// Mitsubishi GX Works2 project: KotelnyaPLC   PLC: FX3U/FX3UC
// Kotelnya

// global labels: Global1
VAR_GLOBAL
  Pw_in_K1 AT D116 : REAL;  (* Давление воды на входе в котел № 1 *)
  TwP_K1 AT D100 : REAL;  (* Температура прямой воды котел № 1 *)
  TwO_K1 AT D102 : REAL;  (* Температура обратной воды котел № 1 *)
  TwP_K2 AT D104 : REAL;  (* Температура прямой воды котел № 2 *)
  TwO_K2 AT D106 : REAL;  (* Температура обратной воды котел № 2 *)
  pusk : BOOL;  (* Переключение вывода данных в градусах "С или "F из блока Fx3U-4AD-PT-ADP *)
  Pw_out_K1 AT D114 : REAL;  (* Давление воды на выходе из котла № 1 *)
  Pw_in_K2 AT D120 : REAL;  (* Давление воды на входе в котел № 2 *)
  Pw_out_K2 AT D118 : REAL;  (* Давление воды на выходе из котла № 2 *)
  TwP AT D108 : REAL;  (* Температура сетевой воды прямой *)
  TwO AT D110 : REAL;  (* Температура сетевой воды обратной *)
  TN_air AT D112 : REAL;  (* Температура наружнего воздуха *)
  F_GAZ AT M144 : BOOL;  (* Флаг активации газового клапана *)
  F_CO_LEVEL2 AT M102 : BOOL;  (* Флаг Активация концентрации по окиси углерода выше 100МГ/М3 Порог 2 *)
  F_CO_LEVEL1 AT M101 : BOOL;  (* Флаг Активация концентрации по окиси углерода выше 20МГ/М3 Порог 1 *)
  F_CH4_LEVEL1 AT M103 : BOOL;  (* Вход Загазованность по метану 0.5% Порог 1 *)
  F_CH4_LEVEL2 AT M104 : BOOL;  (* Вход Загазованность по метану 1% Порог 2 *)
  F_FIRE_RELAY AT M105 : BOOL;  (* Флаг Входа реле пожара *)
  F_HIGH_PRESSURE_GAS AT M146 : BOOL;  (* Флаг Повышение давления газа на вводе *)
  F_LOW_PRESSURE_GAS AT M145 : BOOL;  (* Флаг Понижение давления газа на вводе *)
  F_SB6_SIGNAL_TEST : BOOL;  (* Флаг Тестирование звкового сигнала *)
  F_SB5_SOUND_OFF : BOOL;  (* Флаг Отключение звкового сигнала *)
  F_SA4_SOUND_ON : BOOL;  (* Вход- Переключатель в положении - Звуковой сигнал порога 2 включен *)
  F_SOUND_OFF : BOOL;  (* Флаг Отключение звукового сигнала *)
  F_SOUND : BOOL;  (* Флаг Активация выхода звуковой сигнал *)
  F_LOW_PRESSURE_BACKWATER AT M106 : BOOL;  (* Флаг Понижение давления обратной сетевой воды (унитерм) *)
  F_ALARM_GOR_KOTEL_1 AT M107 : BOOL;  (* Флаг авария Котла 1 *)
  F_ALARM_GOR_KOTEL_2 AT M108 : BOOL;  (* Флаг авария Котла 2 *)
  F_REZERV_PUMP_ON AT M142 : BOOL;  (* Флаг Включился резервный циркуляционный насос. Провод 325 *)
  F_SB1_KOTEL_ON : BOOL;  (* Флаг Кнопка Включения работы Котлов *)
  F_SB2_KOTEL_OFF : BOOL;  (* Флаг Кнопка Выключения работы Котлов *)
  F_SA3_KOTEL_1 : BOOL;  (* Флаг Переключение Котел 1 основной 2 резервный *)
  F_SA3_KOTEL_2 : BOOL;  (* Флаг Переключение Котел 2 основной 1 резервный *)
  F_ROTATION_B_VALVE_COOL AT M201 : BOOL;  (* Флаг Вращение трехходового клапана по часовой стрелке *)
  F_ROTATION_F_VALVE_HEAT AT M202 : BOOL;  (* Флаг Вращение трехходового клапана против часовой стрелки *)
  F_TERMOMETR_95C_KOTEL_1 AT M111 : BOOL;  (* Флаг Термометр манометрический Котел 1. 95С постоянный *)
  F_TERMOMETR_95C_KOTEL_2 AT M112 : BOOL;  (* Флаг Термометр манометрический Котел 2. 95С постоянный *)
  F_SA2_RECIRC_PUMP_1 : BOOL;  (* Флаг. Переключение Рециркуляционный насос 1, Положение Дист *)
  F_SA1_RECIRC_PUMP_1 : BOOL;  (* Флаг. Переключение Рециркуляционный насос 2, Положение Дист *)
  PwP AT D122 : REAL;  (* Давление прямой сетевой воды *)
  PwO AT D124 : REAL;  (* Давление обратной сетевой воды *)
  OP_PwO_ust AT D202 : REAL;  (* ОП Уставка обратного сетевого давления *)
  FB_KOTEL_1 : KOTEL;
  F_KOTEL_1_DOP AT M132 : BOOL;  (* Флаг Котел 1 работает в качестве дополнительного *)
  F_KOTEL_2_DOP AT M134 : BOOL;  (* Флаг Котел 2 работает в качестве дополнительного *)
  F_ALARM_KOTEL_1 AT M135 : BOOL;  (* Флаг Авария Котел 1 *)
  F_ALARM_KOTEL_2 AT M136 : BOOL;  (* Флаг Авария Котел 2 *)
  F_TERMOMETR_90C_KOTEL_1 AT M109 : BOOL;  (* Флаг Термометр манометрический Котел 1. 86С регулируемый *)
  F_TERMOMETR_90C_KOTEL_2 AT M110 : BOOL;  (* Флаг Термометр манометрический Котел 2. 86С регулируемый *)
  OP_PwMAX_ust AT D204 : REAL;  (* Давление воды максимальное Котел *)
  OP_PwMIN_ust AT D206 : REAL;  (* Давление воды минимальное Котел *)
  F_Pdn40_KOTEL_1 AT M113 : BOOL;  (* Флаг Датчик давления в топке ДН-40 Котел 1 *)
  F_Pdn40_KOTEL_2 AT M114 : BOOL;  (* Флаг Датчик давления в топке ДН-40 Котел 2 *)
  OP_Tw80_ust AT D208 : REAL;  (* Панель оператора температура большого горения *)
  OP_Tw86_ust AT D210 : REAL;  (* Панель оператора температура малого горения *)
  F_BURNER_1_KOTEL_1 AT M123 : BOOL;  (* Флаг Горелка 1 Котел 1 *)
  F_BURNER_2_KOTEL_1 AT M124 : BOOL;  (* Флаг Горелка 2 Котел 1 *)
  F_BURNER_1_KOTEL_2 AT M125 : BOOL;  (* Флаг Горелка 1 Котел 2 *)
  F_BURNER_2_KOTEL_2 AT M126 : BOOL;  (* Флаг Горелка 2 Котел 2 *)
  F_CIRC_PUMP_1 AT M140 : BOOL;  (* Флаг Включен циркуляционный насос 1 *)
  F_CIRC_PUMP_2 AT M141 : BOOL;  (* Флаг Включен циркуляционный насос 2 *)
  F_CIRC_PUMP_ON AT M116 : BOOL;  (* Включен циркуляционный насос *)
  F_RECIRC_PUMP_1 AT M127 : BOOL;  (* Флаг активации насоса рециркуляции 1 *)
  F_RECIRC_PUMP_2 AT M128 : BOOL;  (* Флаг активации насоса рециркуляции 2 *)
  OP_RST_ALARM AT M115 : BOOL;  (* Панель оператора Сброс аварии *)
  OP_Tw90_ust AT D212 : REAL;  (* Панель оператора Температура на выходе котла при которой авария *)
  TWO_ust AT D126 : REAL;  (* Температура сетевой воды обратной табличная *)
  OP_GRAPH_N AT D216 : INT;  (* Панель оператора Номер графика нагрева *)
  OP_DAY AT D200 : INT;  (* Панель оператора День *)
  OP_NIGHT AT D201 : INT;  (* Панель оператора Ночь *)
  OP_Tw65_ust AT D214 : REAL;  (* Панель оператора Температура включения рециркуляционного насоса *)
  GRAPH_1 : GRAPH;  (* FBD график определения заданной воды *)
  F_HOUR AT D128 : INT;  (* Час текущий *)
  F_MINUTE AT D129 : INT;  (* Минуты текущие *)
  F_MOTOR_RECIRC_PUMP_1 AT M121 : BOOL;  (* Флаг включен мотор-автомат рециркуляционного насоса 1 *)
  F_MOTOR_RECIRC_PUMP_2 AT M122 : BOOL;  (* Флаг включен мотор-автомат рециркуляционного насоса 2 *)
  F_KOTEL_2 AT M133 : BOOL;  (* Флаг Котел 2 *)
  F_KOTEL_1 AT M131 : BOOL;  (* Флаг Котел 1 *)
  TEMP : BOOL;
  OP_Tw_hist AT D218 : REAL;  (* Панель оператора уставка для горения *)
  F_ALARM_P_KOTEL_1 AT M117 : BOOL;  (* Авария по давлению Котел 1 *)
  FB_KOTEL_2 : KOTEL;
  F_ALARM_P_KOTEL_2 AT M118 : BOOL;  (* Авария по давлению Котел 2 *)
  F_ALARM_T_Water_90_KOTEL_1 AT M119 : BOOL;  (* Авария по температуре 90 градусов Котел 1 *)
  F_ALARM_T_Water_90_KOTEL_2 AT M120 : BOOL;  (* Авария по температуре 90 градусов Котел 2 *)
  TWO_corr AT D220 : INT;  (* Коррекция температуры *)
  F_HL17_LAMP_KOTEL_2 AT M130 : BOOL;  (* Флаг Лампа работы Котла 2 *)
  F_HL16_LAMP_KOTEL_1 AT M129 : BOOL;  (* Флаг Лампа работы Котла 1 *)
  OP_KOTEL_1_2 AT M137 : BOOL;  (* Панель оператора работа котла 1 и 2 одновременно *)
  OP_KOTEL_1_DISABLE AT M501 : BOOL;  (* Панель оператора отключение котла 1 *)
  OP_KOTEL_2_DISABLE AT M502 : BOOL;  (* Панель оператора отключение котла 2 *)
  SCAN_MS : INT;
  TOF_LOW_PRESSURE : TOF;
  OP_ROTATION_F_VALVE_HEAT AT M139 : BOOL;
  OP_ROTATION_F_VALVE_COOL AT M138 : BOOL;
  OP_ALARM_P_sec_KOTEL_1 AT D130 : INT;  (* Время до включения аварии по давлению на котле 1 *)
  OP_ALARM_P_sec_KOTEL_2 AT D131 : INT;  (* Время до включения аварии по давлению на котле 2 *)
  F_ALARM_OUT : BOOL;  (* Флаг Активация аварии общей *)
  OP_ROTATION_POSITION AT D222 : INT;  (* Счет градусов угла поворота трехходового крана *)
  F_RECIRC_PUMP_12 AT M143 : BOOL;  (* Флаг активации рециркуляционных насосов 12 *)
  CIRC_PUMP_1_hour AT D224 : INT;
  CIRC_PUMP_1_min AT D223 : INT;
  CIRC_PUMP_2_min AT D225 : INT;
  CIRC_PUMP_2_hour AT D226 : INT;
  REZERV_PUMP_hour AT D228 : INT;
  REZERV_PUMP_min AT D227 : INT;
  RECIRC_PUMP_12_min AT D229 : INT;
  RECIRC_PUMP_12_hour AT D230 : INT;
  BURNER_1_KOTEL_1_min AT D231 : INT;
  BURNER_1_KOTEL_1_hour AT D232 : INT;
  BURNER_2_KOTEL_1_min AT D233 : INT;
  BURNER_2_KOTEL_1_hour AT D234 : INT;
  BURNER_1_KOTEL_2_min AT D235 : INT;
  BURNER_1_KOTEL_2_hour AT D236 : INT;
  BURNER_2_KOTEL_2_min AT D237 : INT;
  BURNER_2_KOTEL_2_hour AT D238 : INT;
  OP_BIG_FIRE_DOP_1_2 AT D240 : REAL;  (* Панель оператора Уставка включения большого горения и Дополнительного котла *)
  TwO_int AT D133 : INT;  (* Температура воды обратной int *)
  TWO_ust_int AT D132 : INT;  (* Температура обратной воды заданная int *)
  TwP_int AT D134 : INT;  (* Температура прямой воды int *)
  PwP_int AT D135 : INT;  (* Давление прямой сетевой воды, кПа int *)
  PwO_int AT D136 : INT;  (* Давление обратной сетевой воды, кПа int *)
  noi_CIRC_PUMP_1_day_cur AT D137 : INT;
  noi_CIRC_PUMP_1_month_cur AT D138 : INT;
  noi_CIRC_PUMP_1_hour AT D242 : INT;
  noi_CIRC_PUMP_1_day AT D243 : INT;
  noi_CIRC_PUMP_1_month AT D244 : INT;
  noi_CIRC_PUMP_1_month_prev AT D245 : INT;
  noi_CIRC_PUMP_2_day_cur AT D139 : INT;
  noi_CIRC_PUMP_2_month_cur AT D140 : INT;
  noi_CIRC_PUMP_2_hour AT D246 : INT;
  noi_CIRC_PUMP_2_day AT D247 : INT;
  noi_CIRC_PUMP_2_month AT D248 : INT;
  noi_CIRC_PUMP_2_month_prev AT D249 : INT;
  noi_REZERV_PUMP_ON_day_cur AT D141 : INT;
  noi_REZERV_PUMP_ON_month_cur AT D142 : INT;
  noi_REZERV_PUMP_ON_hour AT D250 : INT;
  noi_REZERV_PUMP_ON_day AT D251 : INT;
  noi_REZERV_PUMP_ON_month AT D252 : INT;
  noi_REZERV_PUMP_ON_month_prev AT D253 : INT;
  noi_RECIRC_PUMP_12_day_cur AT D143 : INT;
  noi_RECIRC_PUMP_12_month_cur AT D144 : INT;
  noi_RECIRC_PUMP_12_hour AT D254 : INT;
  noi_RECIRC_PUMP_12_day AT D255 : INT;
  noi_RECIRC_PUMP_12_month AT D256 : INT;
  noi_RECIRC_PUMP_12_month_prev AT D257 : INT;
  noi_BURNER_1_KOTEL_1_day_cur AT D145 : INT;
  noi_BURNER_1_KOTEL_1_month_cur AT D146 : INT;
  noi_BURNER_1_KOTEL_1_hour AT D258 : INT;
  noi_BURNER_1_KOTEL_1_day AT D259 : INT;
  noi_BURNER_1_KOTEL_1_month AT D260 : INT;
  noi_BURNER_1_KOTEL_1_month_prev AT D261 : INT;
  noi_BURNER_2_KOTEL_1_day_cur AT D147 : INT;
  noi_BURNER_2_KOTEL_1_month_cur AT D148 : INT;
  noi_BURNER_2_KOTEL_1_hour AT D262 : INT;
  noi_BURNER_2_KOTEL_1_day AT D263 : INT;
  noi_BURNER_2_KOTEL_1_month AT D264 : INT;
  noi_BURNER_2_KOTEL_1_month_prev AT D265 : INT;
  noi_BURNER_1_KOTEL_2_day_cur AT D149 : INT;
  noi_BURNER_1_KOTEL_2_month_cur AT D150 : INT;
  noi_BURNER_1_KOTEL_2_hour AT D266 : INT;
  noi_BURNER_1_KOTEL_2_day AT D267 : INT;
  noi_BURNER_1_KOTEL_2_month AT D268 : INT;
  noi_BURNER_1_KOTEL_2_month_prev AT D269 : INT;
  noi_BURNER_2_KOTEL_2_day_cur AT D151 : INT;
  noi_BURNER_2_KOTEL_2_month_cur AT D152 : INT;
  noi_BURNER_2_KOTEL_2_hour AT D270 : INT;
  noi_BURNER_2_KOTEL_2_day AT D271 : INT;
  noi_BURNER_2_KOTEL_2_month AT D272 : INT;
  noi_BURNER_2_KOTEL_2_month_prev AT D273 : INT;
  PGAS AT D153 : REAL;  (* Давление газа на вводе *)
  PGAS_int AT D155 : INT;  (* Давление газа на вводе, мБар int *)
  OP_PGAS_min AT D274 : INT;  (* Минимальное давление газа на вводе *)
  OP_PGAS_max AT D275 : INT;  (* Максимальное давление газа на вводе *)
  F_PRESSURE_GAS : BOOL;  (* Флаг Авария по давлению газа на вводе *)
  P_Water_IN_status_KOTEL_1 AT D156 : INT;  (* Состояние давления воды на входе в Котел 1 *)
  P_Water_OUT_status_KOTEL_1 AT D157 : INT;  (* Состояние давления воды на выходе из Котла 1 *)
  P_Water_IN_status_KOTEL_2 AT D158 : INT;  (* Состояние давления воды на входе в Котел 2 *)
  P_Water_OUT_status_KOTEL_2 AT D159 : INT;  (* Состояние давления воды на выходе из Котла 2 *)
END_VAR
VAR_GLOBAL CONSTANT
  RS485_96_8N1 : WORD := 16#1C81;
  RS485_96_8O1 : WORD := 16#1C83;
  RS485_96_8E1 : WORD := 16#1C87;
  RS485_96_8N2 : WORD := 16#1C89;
END_VAR
VAR_GLOBAL
  F_FEEDER_4 AT M147 : BOOL;  (* Флаг питание Фидер 4 *)
  F_FEEDER_26 AT M148 : BOOL;  (* Флаг питание Фидер 26 *)
  VOLTAGE_UA AT D160 : WORD;  (* Напряжение фаза A *)
  VOLTAGE_UB AT D161 : WORD;  (* Напряжение фаза B *)
  VOLTAGE_UC AT D162 : WORD;  (* Напряжение фаза C *)
  VOLTAGE_UAB AT D163 : WORD;  (* Напряжение межфазное AB *)
  VOLTAGE_UBC AT D164 : WORD;  (* Напряжение межфазное BC *)
  VOLTAGE_UCA AT D165 : WORD;  (* Напряжение межфазное CA *)
  VOLTAGE_FREQ AT D166 : WORD;  (* Частота сети, Гц *)
  noi_per_hour_pump_1_MB AT D69 : WORD;
  TwO_ve AT D277 : INT;  (* Температура обратной воды, выше которой разрешен подмес холодной воды *)
  TWO_ust_min AT D276 : INT;  (* Минимальная температура обратной воды заданная *)
  TwO_ve_real : REAL;  (* Температура обратной воды, выше которой разрешен подмес холодной воды *)
  Time_Dop_Kotel_2_min_on AT D168 : INT;  (* Время до включения 2го котла *)
  Time_Dop_Kotel_1_min_on AT D167 : INT;  (* Время до включения 1го котла *)
  F_TIMER_BEFORE_START_KOTEL_1 AT M149 : BOOL;  (* Флаг Индикация таймера до запуска Котла 1 в качестве дополнительного *)
  Time_Dop_Kotel_1_min_off AT D169 : INT;  (* Время до отключения 1го котла *)
  Time_Dop_Kotel_2_min_off AT D170 : INT;  (* Время до отключения 2го котла *)
  F_TIMER_BEFORE_START_KOTEL_2 AT M150 : BOOL;  (* Флаг Индикация таймера до запуска Котла 2 в качестве дополнительного *)
  F_TIMER_BEFORE_STOP_KOTEL_1 AT M151 : BOOL;  (* Флаг Индикация таймера до останова Котла 1 в качестве дополнительного *)
  F_TIMER_BEFORE_STOP_KOTEL_2 AT M152 : BOOL;  (* Флаг Индикация таймера до останова Котла 2 в качестве дополнительного *)
END_VAR

// global labels: DIN
VAR_GLOBAL
  SWT_SA4_SOUND_ON AT X006 : BOOL;  (* Вход- Переключатель в положении - Звуковой сигнал порога 2 включен. Провод 307 *)
  BUT_SB5_SOUND_OFF AT X013 : BOOL;  (* Вход- Отключение звукового сигнала. Провод 312 *)
  BUT_SB6_SIGNAL_TEST AT X014 : BOOL;  (* Вход- Тестирование звукового сигнала. Провод 313 *)
  BUT_SB3_GAZ_ON AT X011 : BOOL;  (* Кнопка включение клапана на вводе газа. NO Контакт 310 *)
  BUT_SB4_GAZ_OFF AT X012 : BOOL;  (* Кнопка выключения клапана на вводе газа. NC Контакт 311 *)
  BUT_SB7_GAZ_TEST : BOOL;  (* Вход Кнопка местного опробования клапана. *)
  DI_CO_LEVEL2 AT X035 : BOOL;  (* Вход Концентрация по окиси углерода выше 100мг/м3 Порог 2. Провод 330 *)
  DI_CO_LEVEL1 AT X034 : BOOL;  (* Вход Концентрация по окиси углерода выше 20мг/м3 Порог 1. Провод 329 *)
  DI_CH4_LEVEL1 AT X036 : BOOL;  (* Вход Загазованность по метану 0.5% Порог 1. Провод 331 *)
  DI_CH4_LEVEL2 AT X037 : BOOL;  (* Вход Загазованность по метану 1% Порог 2. Провод 332 *)
  DI_FIRE_RELAY AT X044 : BOOL;  (* Контакт Реле пожара *)
  DI_K11_ALARM_KOTEL_1 AT X015 : BOOL;  (* Вход авария Котла 1. Провод 314 *)
  DI_K14_ALARM_KOTEL_2 AT X016 : BOOL;  (* Вход авария Котла 2. Провод 315 *)
  DI_REZERV_PUMP_ON AT X027 : BOOL;  (* Вход Включился резервный циркуляционный насос. Провод 324 *)
  BUT_SB1_KOTEL_ON AT X007 : BOOL;  (* Вход Кнопка Включения работы Котлов. Провод 308 *)
  BUT_SB2_KOTEL_OFF AT X010 : BOOL;  (* Вход Кнопка Выключения работы Котлов. Провод 309 *)
  SWT_SA3_KOTEL_1 AT X004 : BOOL;  (* Переключение Котел 1. Провод 305 *)
  SWT_SA3_KOTEL_2 AT X005 : BOOL;  (* Переключение Котел 2. Провод 306 *)
  DI_TERMOMETR_95C_KOTEL_1 AT X020 : BOOL;  (* Вход Термометр манометрический Котел 1. Провод  317 *)
  DI_TERMOMETR_95C_KOTEL_2 AT X024 : BOOL;  (* Вход Термометр манометрический Котел 2. Провод 321 *)
  SWT_SA2_RECIRC_PUMP_1 AT X000 : BOOL;  (* Переключение Рециркуляционный насос 1, Положение Дист. Провод 301 *)
  SWT_SA2_RECIRC_PUMP_2 AT X001 : BOOL;  (* Переключение Рециркуляционный насос 1, Положение Мест. Провод 302 *)
  SWT_SA1_RECIRC_PUMP_1 AT X002 : BOOL;  (* Переключение Рециркуляционный насос 2, Положение Дист. Провод 303 *)
  SWT_SA1_RECIRC_PUMP_2 AT X003 : BOOL;  (* Переключение Рециркуляционный насос 2, Положение Мест. Провод 304 *)
  DI_TERMOMETR_90C_KOTEL_1 AT X017 : BOOL;  (* Вход Термометр манометрический Котел 1. Провод  316 *)
  DI_TERMOMETR_90C_KOTEL_2 AT X023 : BOOL;  (* Вход Термометр манометрический Котел 2. Провод 320 *)
  DI_Pdn40_KOTEL_1 AT X022 : BOOL;  (* Датчик давления в топке ДН-40 Котел 1. Провод 319 *)
  DI_Pdn40_KOTEL_2 AT X026 : BOOL;  (* Датчик давления в топке ДН-40 Котел 2. Провод 323 *)
  DI_CIRC_PUMP_1 AT X030 : BOOL;  (* Вход включился циркуляционный насос 1. Провод 325 *)
  DI_CIRC_PUMP_2 AT X031 : BOOL;  (* Вход включился циркуляционный насос 2. Провод 326 *)
  DI_MOTOR_RECIRC_PUMP_1 AT X032 : BOOL;  (* Вход включен мотор-автомат рециркуляционного насоса 1. Провод 327 *)
  DI_MOTOR_RECIRC_PUMP_2 AT X033 : BOOL;  (* Вход включен мотор-автомат рециркуляционного насоса 2. Провод 328 *)
  DI_FEEDER_4 AT X042 : BOOL;  (* Вход Питание Фидер 4. Провод 335 *)
  DI_FEEDER_26 AT X043 : BOOL;  (* Вход Питание Фидер 26. Провод 336 *)
  DI_P_DIF_ALARM AT X045 : BOOL;  (* Вход Авария по перепаду давления дифманометра НО контакт. Провод 338 *)
END_VAR

// global labels: DOUT
VAR_GLOBAL
  DO_ROTATION_B_VALVE AT Y001 : BOOL;  (* Резервный насос 30 кВт. Провод 403 *)
  DO_R4_SOUND AT Y003 : BOOL;  (* Выход звуковая сирена. Провод 404 *)
  DO_ROTATION_F_VALVE AT Y002 : BOOL;  (* Котел 2. Провод 402 *)
  DO_LAMP_CH4_LEVEL1 AT Y006 : BOOL;  (* Загазованность по "СН" порог 1. Провод 407 *)
  DO_LAMP_CO_LEVEL2 AT Y007 : BOOL;  (* Концентрация по "СO" порог 2. Провод 408 *)
  DO_LAMP_CO_LEVEL1 AT Y010 : BOOL;  (* Концентрация по "СO" порог 1. Провод 409 *)
  DO_HL5_LAMP_PRESSURE_GAZ_LOW AT Y011 : BOOL;  (* Давление газа низкое. Провод 410 *)
  DO_HL6_LAMP_PRESSURE_GAZ_HIGH AT Y012 : BOOL;  (* Давление газа высокое. Провод 411 *)
  DO_LAMP_CH4_LEVEL2 AT Y021 : BOOL;  (* Загазованность по "СН4" порог 2. Провод 418 *)
  DO_HL14_LAMP_PUMP_RECIRCULATON_2 AT Y022 : BOOL;  (* Насос рециркуляции № 2. Провод 419 *)
  DO_HL15_LAMP_PUMP_RECIRCULATON_1 AT Y023 : BOOL;  (* Насос рециркуляции № 1. Провод 420 *)
  DO_HL16_LAMP_KOTEL_1 AT Y024 : BOOL;  (* Лампа. Котел № 1. Провод 421 *)
  DO_HL17_LAMP_KOTEL_2 AT Y025 : BOOL;  (* Лампа Котел № 2. Провод 422 *)
  DO_HL7_R7_LAMP_GAZ_ON AT Y013 : BOOL;  (* Выход Лампа газовый клапан включен и Активация реле R7 включение газового клапана *)
  DO_HL12_LAMP_GAZ_OFF AT Y020 : BOOL;  (* Выход Лампа газовый клапан выключен. Провод 417 *)
  DO_LAMP_LOW_PRESSURE_BACKWATER AT Y015 : BOOL;  (* Выход лампа Давления обратной сетевой воды низкое (унитерм). Контакт 414 *)
  DO_LAMP_ALARM_KOTEL_1 AT Y017 : BOOL;  (* Выход Лампа Авария котел 1. Провод 416 *)
  DO_LAMP_ALARM_KOTEL_2 AT Y016 : BOOL;  (* Выход Лампа Авария котел 2. Провод 415 *)
  DO_LAMP_REZERV_PUMP_ON AT Y014 : BOOL;  (* Выход лампа Включился резервный циркуляционный насос. Провод 413 *)
  DO_PUMP_RECIRCULATION_1 AT Y004 : BOOL;  (* Рециркуляционный насос 1. Провод 405 *)
  DO_PUMP_RECIRCULATION_2 AT Y005 : BOOL;  (* Рециркуляционный насос 2. Провод 406 *)
  DO_BURNER_1_KOTEL_1 AT Y026 : BOOL;  (* Выход Горелка 1 Котел 1. Провод 423 *)
  DO_BURNER_2_KOTEL_1 AT Y027 : BOOL;  (* Выход Горелка 2 Котел 1. Провод 424 *)
  DO_BURNER_1_KOTEL_2 AT Y022 : BOOL;  (* Выход Горелка 1 Котел 2. Провод 425 *)
  DO_BURNER_2_KOTEL_2 AT Y023 : BOOL;  (* Выход Горелка 2 Котел 2. Провод 426 *)
  DO_ALARM_OUT AT Y000 : BOOL;  (* Выход Активация аварии общей *)
  EXT_ALARM_GOR_1 AT Y040 : BOOL;  (* Выход сигнализация Авария горелки 1 *)
  EXT_ALARM_GOR_2 AT Y042 : BOOL;  (* Выход сигнализация Авария горелки 2 *)
  EXT_ALARM_KOTEL_1 AT Y041 : BOOL;  (* Выход сигнализация Авария Котел 1 *)
  EXT_ALARM_KOTEL_2 AT Y043 : BOOL;  (* Выход сигнализация Авария Котел 2 *)
  EXT_ALARM_GAZ_OFF AT Y044 : BOOL;  (* Выход сигнализация Авария по закрытии газового клапана *)
  EXT_ALARM_P_DIF_ALARM AT Y045 : BOOL;  (* Выход сигнализация Авария по перепаду давления дифманометра *)
  EXT_ALARM_LOW_PRESSURE_WATER AT Y046 : BOOL;  (* Выход по низкому давлению воды *)
  EXT_ALARM_NONE_VOLTAGE AT Y047 : BOOL;  (* Выход сигнализация Отсутствие сети по 4 и 26 фидеру *)
END_VAR

// global labels: Water
VAR_GLOBAL
  WATER_LEVEL AT D50 : WORD;  (* Уровень воды в баке водоподготовки *)
  PRESSURE_BEFORE_FILTER AT D51 : WORD;  (* Давление до фильтра *)
  PRESSURE_AFTER_FILTER AT D52 : WORD;  (* Давление после фильтра *)
  CAPACITY_HOUR_MB AT D53 : WORD;
  CAPACITY_DAY_MB AT D54 : WORD;
  CAPACITY_MONTH_MB AT D55 : WORD;
  CAPACITY_HOUR_cur_MB AT D56 : WORD;
  CAPACITY_DAY_cur_MB AT D57 : WORD;
  CAPACITY_MONTH_cur_MB AT D58 : WORD;
  NOI_DAY_PUMP_1_cur_MB AT D59 : WORD;
  NOI_MONTH_PUMP_1_cur_MB AT D60 : WORD;
  NOI_DAY_PUMP_2_cur_MB AT D61 : WORD;
  NOI_MONTH_PUMP_2_cur_MB AT D62 : WORD;
  number_of_inclusions_pump_1_MB AT D63 : WORD;
  number_of_inclusions_pump_2_MB AT D65 : WORD;
  noi_pump_1_cur_MB AT D67 : WORD;
  noi_pump_2_cur_MB AT D68 : WORD;
  noi_per_hour_pump_2_MB AT D70 : WORD;
  noi_per_day_pump_1_MB AT D71 : WORD;
  noi_per_day_pump_2_MB AT D72 : WORD;
  noi_per_month_pump_1_MB AT D73 : WORD;
  noi_per_month_pump_2_MB AT D74 : WORD;
  F_FILLING_VALVE_MB AT M75 : BOOL;
  F_DUMP_VALVE_MB AT M76 : BOOL;
  F_PUMP_1_MB AT M77 : BOOL;
  F_PUMP_2_MB AT M78 : BOOL;
  OP_PUMP_12_MB AT M79 : BOOL;
END_VAR

// task Task_01 (event TRUE, interval 0, priority 31): AIN_FBD, COUNTERS, MAIN, EXT_ALARM, FX3UModbusRTUMaster_PRG, VOLTAGE
// user libraries (not included): AnalogFX_V100, FX3UModbusRTUMaster_V100

PROGRAM MAIN
VAR
  TON_VALVE_1 : TON;
  TOF_VALVE_1 : TOF;
  TOF_VALVE_2 : TOF;
  TON_VALVE_2 : TON;
  F_ROTATION_F_VALVE_HEAT_CNT : INT;
  F_ROTATION_F_VALVE_HEAT_ENABLE : BOOL;
  F_ROTATION_F_VALVE_COOL_CNT : INT;
  F_ROTATION_F_VALVE_COOL_ENABLE : BOOL;
  TOF_CIRC_PUMP_ON : TOF;
  TOF_LOW_PRESSURE_M8002 : TOF;
  TON_GAS_HIGH : TON;
  TON_GAS_LOW : TON;
  TOF_RECIRC_PUMP_1 : TOF;
  TOF_RECIRC_PUMP_2 : TOF;
END_VAR
(* structured ladder/FBD written out as ST: instructions are called as NAME(EN, inputs, outputs); _pN, _eN, _tN stand for wires *)
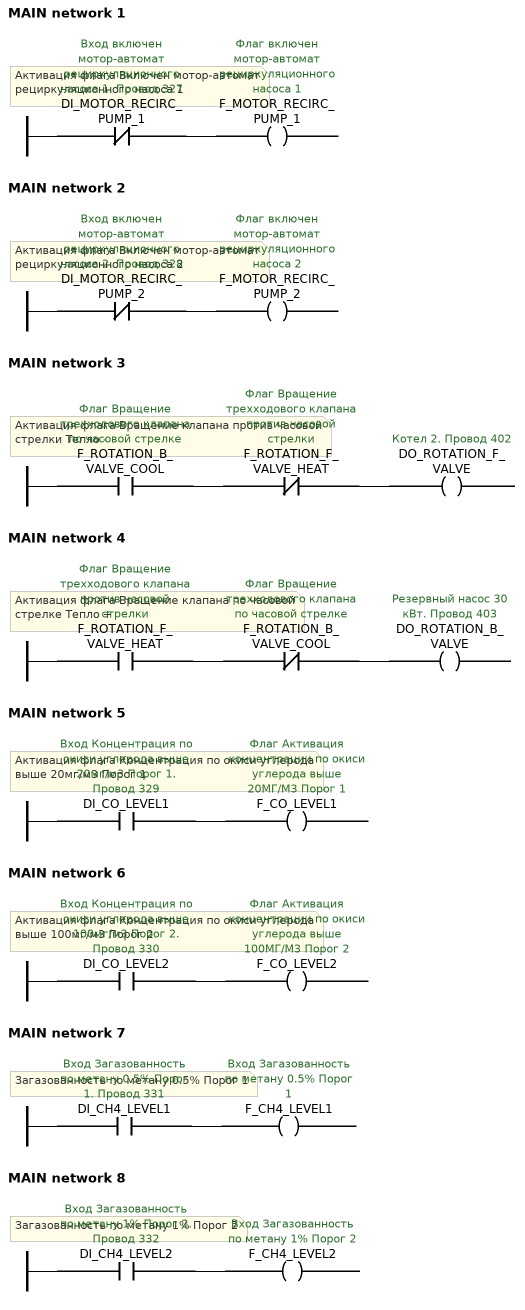
(* network 1 *)
(* Активация флага Включен мотор-автомат рециркуляционного насоса 1 *)
F_MOTOR_RECIRC_PUMP_1 := NOT DI_MOTOR_RECIRC_PUMP_1;
(* network 2 *)
(* Активация флага Включен мотор-автомат рециркуляционного насоса 2 *)
F_MOTOR_RECIRC_PUMP_2 := NOT DI_MOTOR_RECIRC_PUMP_2;
(* network 3 *)
(* Активация флага Вращение клапана против часовой стрелки Тепло - *)
DO_ROTATION_F_VALVE := F_ROTATION_B_VALVE_COOL AND NOT F_ROTATION_F_VALVE_HEAT;
(* network 4 *)
(* Активация флага Вращение клапана по часовой стрелке Тепло + *)
DO_ROTATION_B_VALVE := F_ROTATION_F_VALVE_HEAT AND NOT F_ROTATION_B_VALVE_COOL;
(* network 5 *)
(* Активация флага Концентрация по окиси углерода выше 20мг/м3 Порог 1 *)
F_CO_LEVEL1 := DI_CO_LEVEL1;
(* network 6 *)
(* Активация флага Концентрация по окиси углерода выше 100мг/м3 Порог 2 *)
F_CO_LEVEL2 := DI_CO_LEVEL2;
(* network 7 *)
(* Загазованность по метану 0.5% Порог 1 *)
F_CH4_LEVEL1 := DI_CH4_LEVEL1;
(* network 8 *)
(* Загазованность по метану 1% Порог 2 *)
F_CH4_LEVEL2 := DI_CH4_LEVEL2;
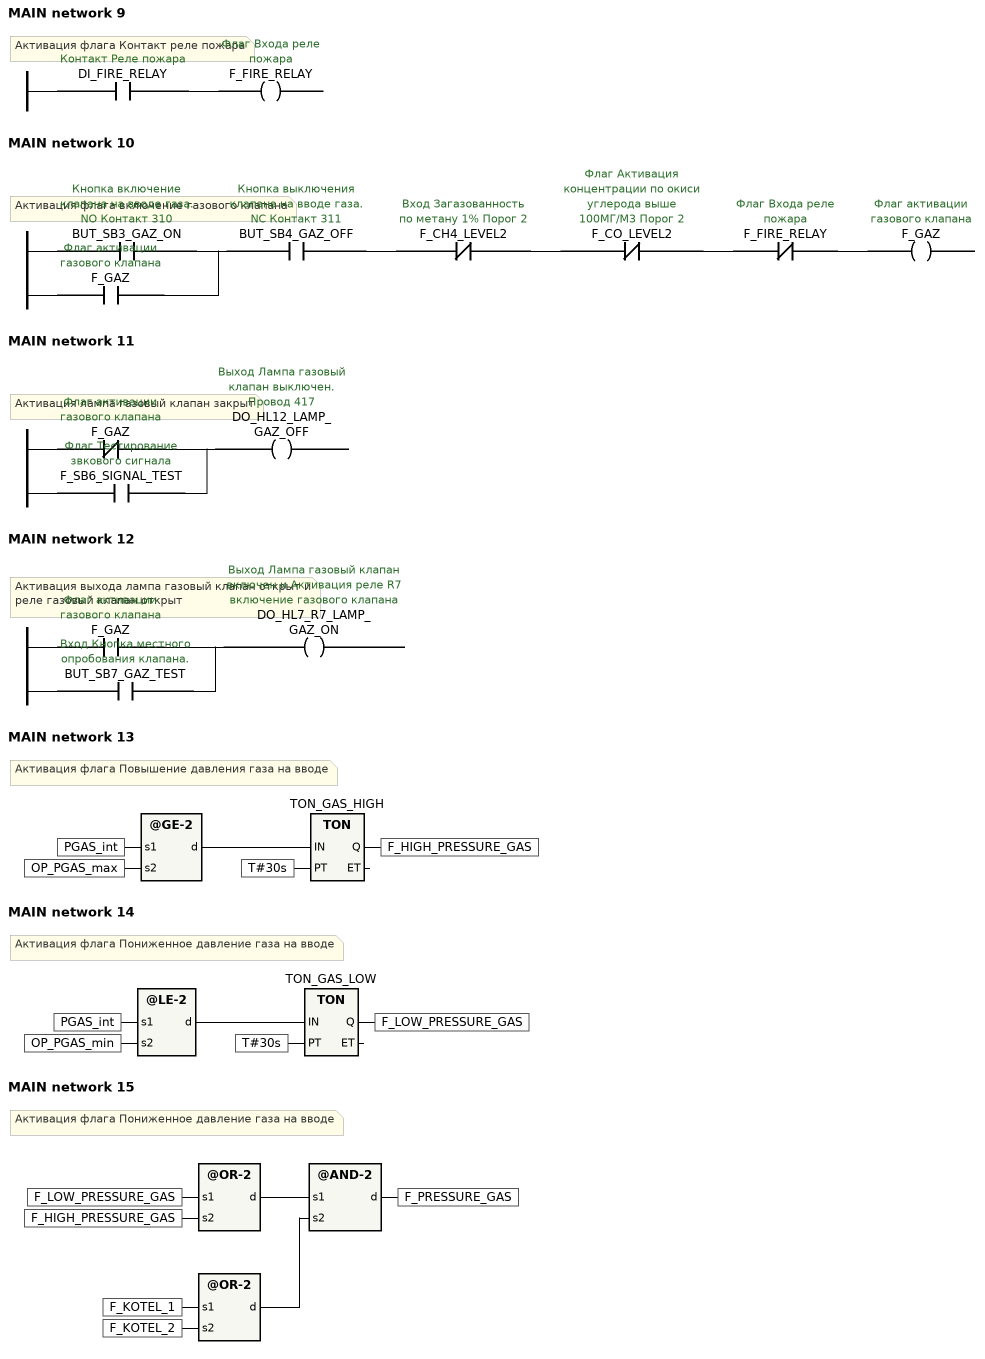
(* network 9 *)
(* Активация флага Контакт реле пожара *)
F_FIRE_RELAY := DI_FIRE_RELAY;
(* network 10 *)
(* Активация флага включение газового клапана *)
F_GAZ := ((((BUT_SB3_GAZ_ON OR F_GAZ) AND BUT_SB4_GAZ_OFF) AND NOT F_CH4_LEVEL2) AND NOT F_CO_LEVEL2) AND NOT F_FIRE_RELAY;
(* network 11 *)
(* Активация лампа газовый клапан закрыт *)
DO_HL12_LAMP_GAZ_OFF := (NOT F_GAZ) OR F_SB6_SIGNAL_TEST;
(* network 12 *)
(* Активация выхода лампа газовый клапан открыт и реле газовый клапан открыт *)
DO_HL7_R7_LAMP_GAZ_ON := F_GAZ OR BUT_SB7_GAZ_TEST;
(* network 13 *)
(* Активация флага Повышение давления газа на вводе *)
TON_GAS_HIGH(IN := @GE-2(PGAS_int, OP_PGAS_max), PT := T#30s, Q => F_HIGH_PRESSURE_GAS);
(* network 14 *)
(* Активация флага Пониженное давление газа на вводе *)
TON_GAS_LOW(IN := @LE-2(PGAS_int, OP_PGAS_min), PT := T#30s, Q => F_LOW_PRESSURE_GAS);
(* network 15 *)
(* Активация флага Пониженное давление газа на вводе *)
F_PRESSURE_GAS := @AND-2(@OR-2(F_LOW_PRESSURE_GAS, F_HIGH_PRESSURE_GAS), @OR-2(F_KOTEL_1, F_KOTEL_2));
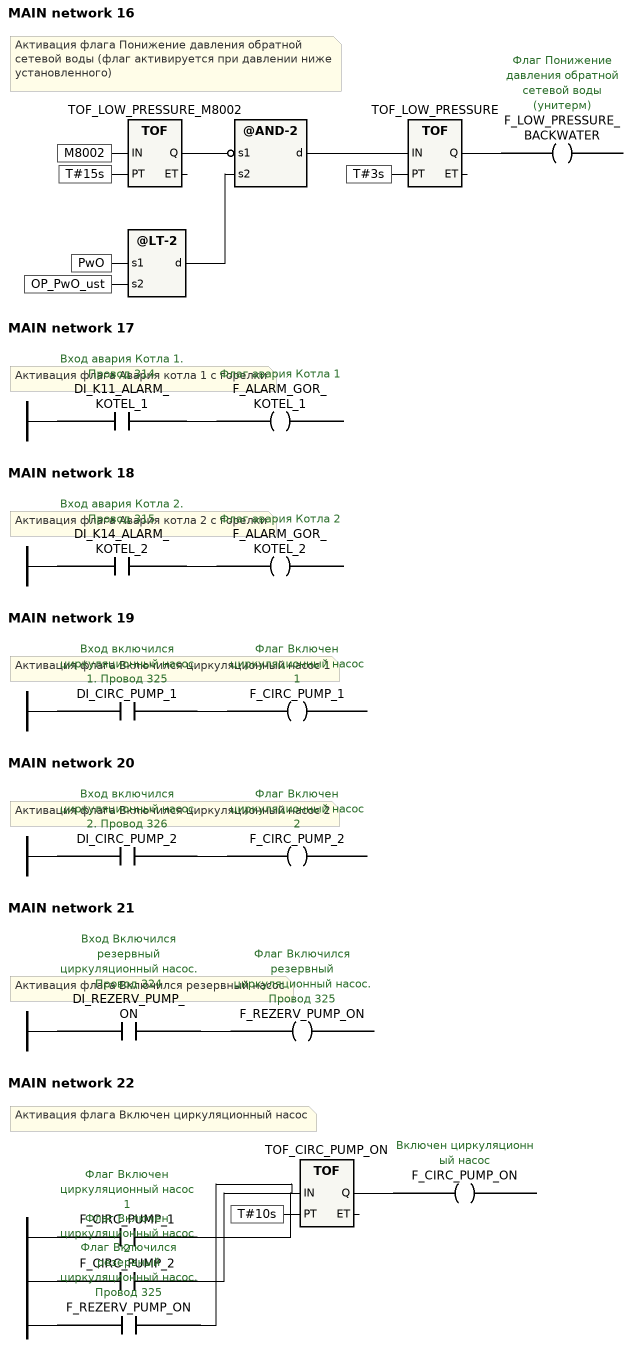
(* network 16 *)
(* Активация флага Понижение давления обратной сетевой воды (флаг активируется при давлении ниже установленного) *)
TOF_LOW_PRESSURE_M8002(IN := M8002, PT := T#15s);
TOF_LOW_PRESSURE(IN := @AND-2(NOT TOF_LOW_PRESSURE_M8002.Q, @LT-2(PwO, OP_PwO_ust)), PT := T#3s);
F_LOW_PRESSURE_BACKWATER := TOF_LOW_PRESSURE.Q;
(* network 17 *)
(* Активация флага Авария котла 1 с горелки *)
F_ALARM_GOR_KOTEL_1 := DI_K11_ALARM_KOTEL_1;
(* network 18 *)
(* Активация флага Авария котла 2 с горелки *)
F_ALARM_GOR_KOTEL_2 := DI_K14_ALARM_KOTEL_2;
(* network 19 *)
(* Активация флага Включился циркуляционный насос 1 *)
F_CIRC_PUMP_1 := DI_CIRC_PUMP_1;
(* network 20 *)
(* Активация флага Включился циркуляционный насос 2 *)
F_CIRC_PUMP_2 := DI_CIRC_PUMP_2;
(* network 21 *)
(* Активация флага Включился резервный насос *)
F_REZERV_PUMP_ON := DI_REZERV_PUMP_ON;
(* network 22 *)
(* Активация флага Включен циркуляционный насос *)
TOF_CIRC_PUMP_ON(IN := F_CIRC_PUMP_1 OR F_CIRC_PUMP_2 OR F_REZERV_PUMP_ON, PT := T#10s);
F_CIRC_PUMP_ON := TOF_CIRC_PUMP_ON.Q;
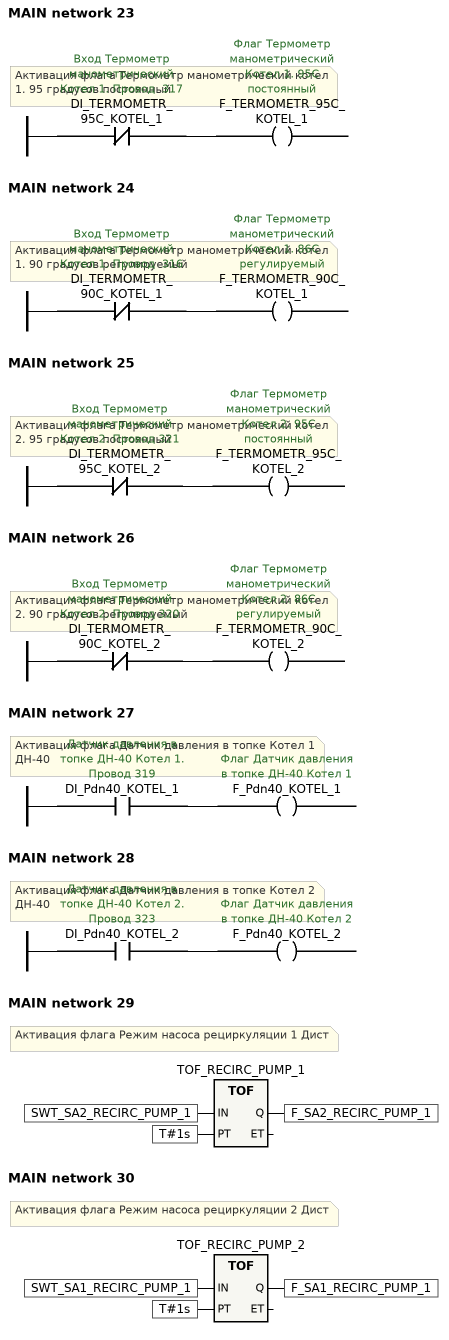
(* network 23 *)
(* Активация флага Термометр манометрический котел 1. 95 градусов постоянный *)
F_TERMOMETR_95C_KOTEL_1 := NOT DI_TERMOMETR_95C_KOTEL_1;
(* network 24 *)
(* Активация флага Термометр манометрический котел 1. 90 градусов регулируемый *)
F_TERMOMETR_90C_KOTEL_1 := NOT DI_TERMOMETR_90C_KOTEL_1;
(* network 25 *)
(* Активация флага Термометр манометрический котел 2. 95 градусов постоянный *)
F_TERMOMETR_95C_KOTEL_2 := NOT DI_TERMOMETR_95C_KOTEL_2;
(* network 26 *)
(* Активация флага Термометр манометрический котел 2. 90 градусов регулируемый *)
F_TERMOMETR_90C_KOTEL_2 := NOT DI_TERMOMETR_90C_KOTEL_2;
(* network 27 *)
(* Активация флага Датчик давления в топке Котел 1 ДН-40 *)
F_Pdn40_KOTEL_1 := DI_Pdn40_KOTEL_1;
(* network 28 *)
(* Активация флага Датчик давления в топке Котел 2 ДН-40 *)
F_Pdn40_KOTEL_2 := DI_Pdn40_KOTEL_2;
(* network 29 *)
(* Активация флага Режим насоса рециркуляции 1 Дист *)
TOF_RECIRC_PUMP_1(IN := SWT_SA2_RECIRC_PUMP_1, PT := T#1s, Q => F_SA2_RECIRC_PUMP_1);
(* network 30 *)
(* Активация флага Режим насоса рециркуляции 2 Дист *)
TOF_RECIRC_PUMP_2(IN := SWT_SA1_RECIRC_PUMP_1, PT := T#1s, Q => F_SA1_RECIRC_PUMP_1);
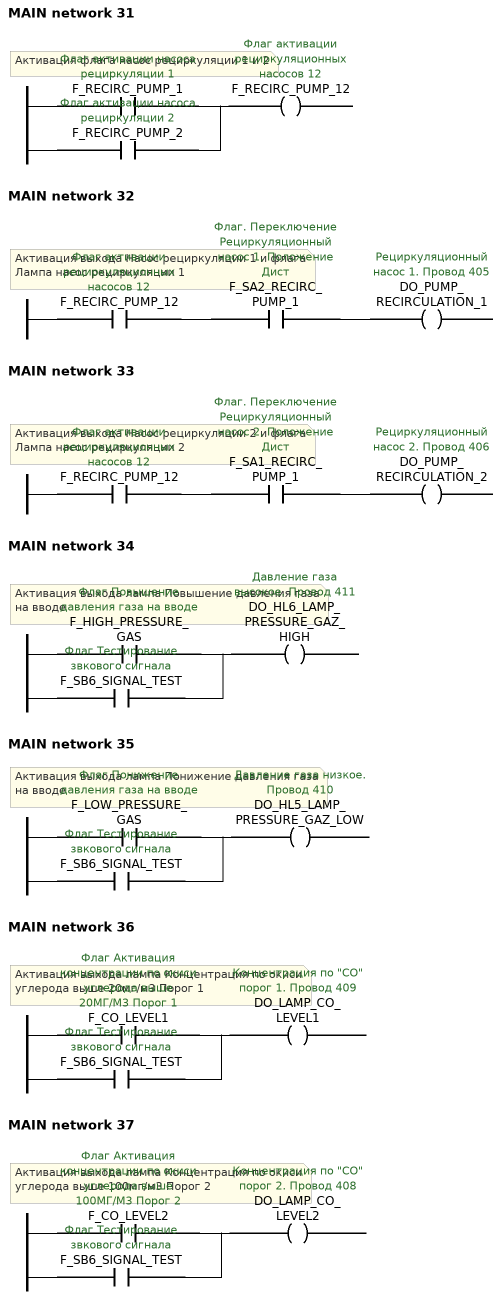
(* network 31 *)
(* Активация флага насос рециркуляции 1 и 2 *)
F_RECIRC_PUMP_12 := F_RECIRC_PUMP_1 OR F_RECIRC_PUMP_2;
(* network 32 *)
(* Активация выхода Насос рециркуляции 1 и флага Лампа насос рециркуляции 1 *)
DO_PUMP_RECIRCULATION_1 := F_RECIRC_PUMP_12 AND F_SA2_RECIRC_PUMP_1;
(* network 33 *)
(* Активация выхода Насос рециркуляции 2 и флага Лампа насос рециркуляции 2 *)
DO_PUMP_RECIRCULATION_2 := F_RECIRC_PUMP_12 AND F_SA1_RECIRC_PUMP_1;
(* network 34 *)
(* Активация выхода лампа Повышение давления газа на вводе *)
DO_HL6_LAMP_PRESSURE_GAZ_HIGH := F_HIGH_PRESSURE_GAS OR F_SB6_SIGNAL_TEST;
(* network 35 *)
(* Активация выхода лампа Понижение давления газа на вводе *)
DO_HL5_LAMP_PRESSURE_GAZ_LOW := F_LOW_PRESSURE_GAS OR F_SB6_SIGNAL_TEST;
(* network 36 *)
(* Активация выхода лампа Концентрация по окиси углерода выше 20мг/м3 Порог 1 *)
DO_LAMP_CO_LEVEL1 := F_CO_LEVEL1 OR F_SB6_SIGNAL_TEST;
(* network 37 *)
(* Активация выхода лампа Концентрация по окиси углерода выше 100мг/м3 Порог 2 *)
DO_LAMP_CO_LEVEL2 := F_CO_LEVEL2 OR F_SB6_SIGNAL_TEST;